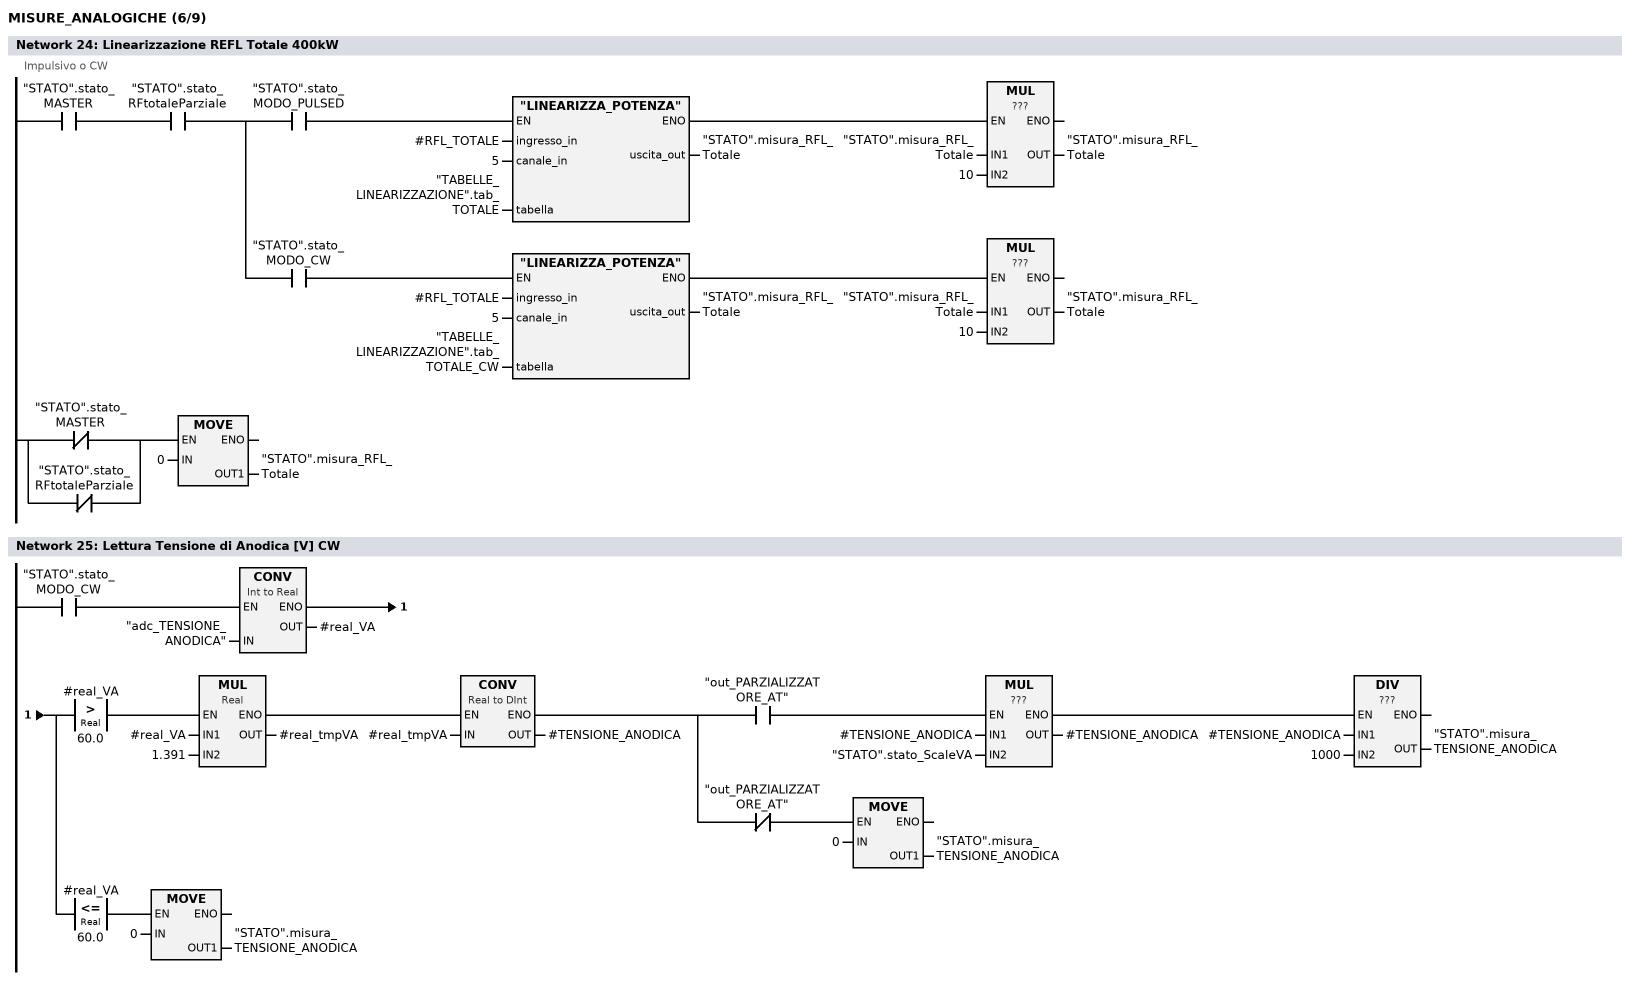
   RUNG wire#powerrail
      Contact( "STATO".stato_MASTER )
      Contact( "STATO".stato_RFtotaleParziale )
      wire#w1
      Contact( "STATO".stato_MODO_PULSED )
      "LINEARIZZA_POTENZA"(ingresso_in := #RFL_TOTALE, canale_in := 5, tabella := "TABELLE_LINEARIZZAZIONE".tab_TOTALE, uscita_out => "STATO".misura_RFL_Totale)
      { S7_Templates := "SrcType := ???" } Mul(in1 := "STATO".misura_RFL_Totale, in2 := 10, out => "STATO".misura_RFL_Totale)
   END_RUNG
   RUNG wire#w1
      Contact( "STATO".stato_MODO_CW )
      "LINEARIZZA_POTENZA"(ingresso_in := #RFL_TOTALE, canale_in := 5, tabella := "TABELLE_LINEARIZZAZIONE".tab_TOTALE_CW, uscita_out => "STATO".misura_RFL_Totale)
      { S7_Templates := "SrcType := ???" } Mul(in1 := "STATO".misura_RFL_Totale, in2 := 10, out => "STATO".misura_RFL_Totale)
   END_RUNG
   RUNG wire#powerrail
      I_Contact( "STATO".stato_MASTER )
      wire#w2
      Move(in := 0, out1 => "STATO".misura_RFL_Totale)
   END_RUNG
   RUNG wire#powerrail
      I_Contact( "STATO".stato_RFtotaleParziale )
   END_RUNG wire#w2
   // the same network as SCL:
   #_w1 := "STATO".stato_MASTER AND "STATO".stato_RFtotaleParziale;
   "LINEARIZZA_POTENZA"(EN := #_w1 AND "STATO".stato_MODO_PULSED,
                        ingresso_in := #RFL_TOTALE,
                        canale_in := 5,
                        tabella := "TABELLE_LINEARIZZAZIONE".tab_TOTALE,
                        uscita_out => "STATO".misura_RFL_Totale,
                        ENO => #_w2);
   IF #_w2 THEN "STATO".misura_RFL_Totale := "STATO".misura_RFL_Totale * 10; END_IF;
   "LINEARIZZA_POTENZA"(EN := #_w1 AND "STATO".stato_MODO_CW,
                        ingresso_in := #RFL_TOTALE,
                        canale_in := 5,
                        tabella := "TABELLE_LINEARIZZAZIONE".tab_TOTALE_CW,
                        uscita_out => "STATO".misura_RFL_Totale,
                        ENO => #_w3);
   IF #_w3 THEN "STATO".misura_RFL_Totale := "STATO".misura_RFL_Totale * 10; END_IF;
   IF NOT "STATO".stato_MASTER OR NOT "STATO".stato_RFtotaleParziale THEN
       "STATO".misura_RFL_Totale := 0;
   END_IF;
END_REGION

REGION Network 25: Lettura Tensione di Anodica [V] CW
   RUNG wire#powerrail
      Contact( "STATO".stato_MODO_CW )
      { S7_Templates := "[SrcType := Int, DestType := Real]" } Convert(in := "adc_TENSIONE_ANODICA", out => #real_VA)
      wire#w1
      { S7_Templates := "SrcType := Real" } GT_Contact(in1 := #real_VA, in2 := 60.0)
      { S7_Templates := "SrcType := Real" } Mul(in1 := #real_VA, in2 := 1.391, out => #real_tmpVA)
      { S7_Templates := "[SrcType := Real, DestType := DInt]" } Convert(in := #real_tmpVA, out => #TENSIONE_ANODICA)
      wire#w2
      Contact( "out_PARZIALIZZATORE_AT" )
      { S7_Templates := "SrcType := ???" } Mul(in1 := #TENSIONE_ANODICA, in2 := "STATO".stato_ScaleVA, out => #TENSIONE_ANODICA)
      { S7_Templates := "SrcType := ???" } Div(in1 := #TENSIONE_ANODICA, in2 := 1000, out => "STATO".misura_TENSIONE_ANODICA)
   END_RUNG
   RUNG wire#w2
      I_Contact( "out_PARZIALIZZATORE_AT" )
      Move(in := 0, out1 => "STATO".misura_TENSIONE_ANODICA)
   END_RUNG
   RUNG wire#w1
      { S7_Templates := "SrcType := Real" } LE_Contact(in1 := #real_VA, in2 := 60.0)
      Move(in := 0, out1 => "STATO".misura_TENSIONE_ANODICA)
   END_RUNG
   // the same network as SCL:
   IF "STATO".stato_MODO_CW THEN #real_VA := INT_TO_REAL("adc_TENSIONE_ANODICA"); END_IF;
   #_w1 := "STATO".stato_MODO_CW AND (#real_VA > 60.0);
   IF #_w1 THEN
       #real_tmpVA := #real_VA * 1.391;
       #TENSIONE_ANODICA := REAL_TO_DINT(#real_tmpVA);
   END_IF;
   IF #_w1 AND "out_PARZIALIZZATORE_AT" THEN
       #TENSIONE_ANODICA := #TENSIONE_ANODICA * "STATO".stato_ScaleVA;
       "STATO".misura_TENSIONE_ANODICA := #TENSIONE_ANODICA / 1000;
   END_IF;
   IF #_w1 AND NOT "out_PARZIALIZZATORE_AT" THEN "STATO".misura_TENSIONE_ANODICA := 0; END_IF;
   IF "STATO".stato_MODO_CW AND (#real_VA <= 60.0) THEN "STATO".misura_TENSIONE_ANODICA := 0; END_IF;
END_REGION

REGION Network 26: Lettura Tensione di Anodica [V] PULSED
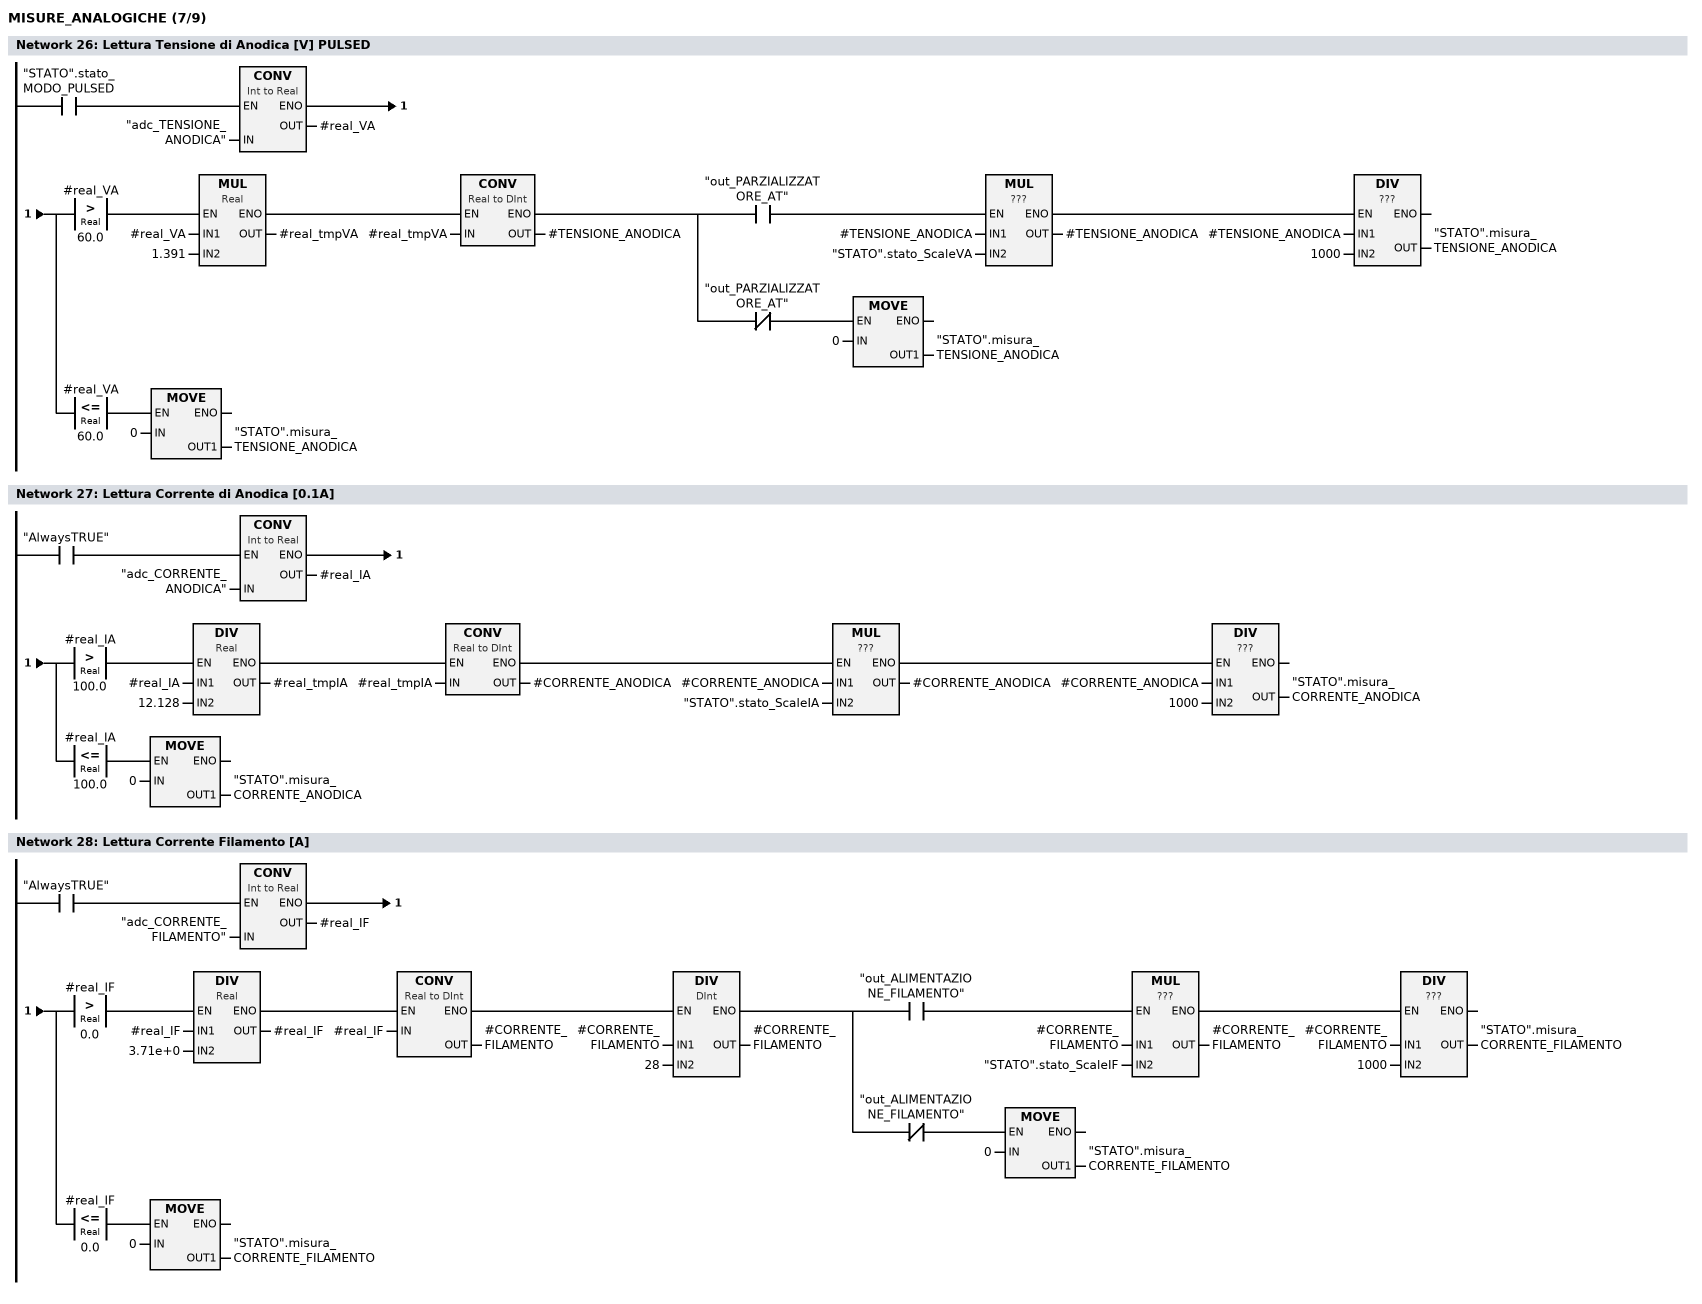
   RUNG wire#powerrail
      Contact( "STATO".stato_MODO_PULSED )
      { S7_Templates := "[SrcType := Int, DestType := Real]" } Convert(in := "adc_TENSIONE_ANODICA", out => #real_VA)
      wire#w1
      { S7_Templates := "SrcType := Real" } GT_Contact(in1 := #real_VA, in2 := 60.0)
      { S7_Templates := "SrcType := Real" } Mul(in1 := #real_VA, in2 := 1.391, out => #real_tmpVA)
      { S7_Templates := "[SrcType := Real, DestType := DInt]" } Convert(in := #real_tmpVA, out => #TENSIONE_ANODICA)
      wire#w2
      Contact( "out_PARZIALIZZATORE_AT" )
      { S7_Templates := "SrcType := ???" } Mul(in1 := #TENSIONE_ANODICA, in2 := "STATO".stato_ScaleVA, out => #TENSIONE_ANODICA)
      { S7_Templates := "SrcType := ???" } Div(in1 := #TENSIONE_ANODICA, in2 := 1000, out => "STATO".misura_TENSIONE_ANODICA)
   END_RUNG
   RUNG wire#w2
      I_Contact( "out_PARZIALIZZATORE_AT" )
      Move(in := 0, out1 => "STATO".misura_TENSIONE_ANODICA)
   END_RUNG
   RUNG wire#w1
      { S7_Templates := "SrcType := Real" } LE_Contact(in1 := #real_VA, in2 := 60.0)
      Move(in := 0, out1 => "STATO".misura_TENSIONE_ANODICA)
   END_RUNG
   // the same network as SCL:
   IF "STATO".stato_MODO_PULSED THEN #real_VA := INT_TO_REAL("adc_TENSIONE_ANODICA"); END_IF;
   #_w1 := "STATO".stato_MODO_PULSED AND (#real_VA > 60.0);
   IF #_w1 THEN
       #real_tmpVA := #real_VA * 1.391;
       #TENSIONE_ANODICA := REAL_TO_DINT(#real_tmpVA);
   END_IF;
   IF #_w1 AND "out_PARZIALIZZATORE_AT" THEN
       #TENSIONE_ANODICA := #TENSIONE_ANODICA * "STATO".stato_ScaleVA;
       "STATO".misura_TENSIONE_ANODICA := #TENSIONE_ANODICA / 1000;
   END_IF;
   IF #_w1 AND NOT "out_PARZIALIZZATORE_AT" THEN "STATO".misura_TENSIONE_ANODICA := 0; END_IF;
   IF "STATO".stato_MODO_PULSED AND (#real_VA <= 60.0) THEN "STATO".misura_TENSIONE_ANODICA := 0; END_IF;
END_REGION

REGION Network 27: Lettura Corrente di Anodica [0.1A]
   RUNG wire#powerrail
      Contact( "AlwaysTRUE" )
      { S7_Templates := "[SrcType := Int, DestType := Real]" } Convert(in := "adc_CORRENTE_ANODICA", out => #real_IA)
      wire#w1
      { S7_Templates := "SrcType := Real" } GT_Contact(in1 := #real_IA, in2 := 100.0)
      { S7_Templates := "SrcType := Real" } Div(in1 := #real_IA, in2 := 12.128, out => #real_tmpIA)
      { S7_Templates := "[SrcType := Real, DestType := DInt]" } Convert(in := #real_tmpIA, out => #CORRENTE_ANODICA)
      { S7_Templates := "SrcType := ???" } Mul(in1 := #CORRENTE_ANODICA, in2 := "STATO".stato_ScaleIA, out => #CORRENTE_ANODICA)
      { S7_Templates := "SrcType := ???" } Div(in1 := #CORRENTE_ANODICA, in2 := 1000, out => "STATO".misura_CORRENTE_ANODICA)
   END_RUNG
   RUNG wire#w1
      { S7_Templates := "SrcType := Real" } LE_Contact(in1 := #real_IA, in2 := 100.0)
      Move(in := 0, out1 => "STATO".misura_CORRENTE_ANODICA)
   END_RUNG
   // the same network as SCL:
   IF "AlwaysTRUE" THEN #real_IA := INT_TO_REAL("adc_CORRENTE_ANODICA"); END_IF;
   IF "AlwaysTRUE" AND (#real_IA > 100.0) THEN
       #real_tmpIA := #real_IA / 12.128;
       #CORRENTE_ANODICA := REAL_TO_DINT(#real_tmpIA);
       #CORRENTE_ANODICA := #CORRENTE_ANODICA * "STATO".stato_ScaleIA;
       "STATO".misura_CORRENTE_ANODICA := #CORRENTE_ANODICA / 1000;
   END_IF;
   IF "AlwaysTRUE" AND (#real_IA <= 100.0) THEN "STATO".misura_CORRENTE_ANODICA := 0; END_IF;
END_REGION

REGION Network 28: Lettura Corrente Filamento [A]
   RUNG wire#powerrail
      Contact( "AlwaysTRUE" )
      { S7_Templates := "[SrcType := Int, DestType := Real]" } Convert(in := "adc_CORRENTE_FILAMENTO", out => #real_IF)
      wire#w1
      { S7_Templates := "SrcType := Real" } GT_Contact(in1 := #real_IF, in2 := 0.0)
      { S7_Templates := "SrcType := Real" } Div(in1 := #real_IF, in2 := 3.71e+0, out => #real_IF)
      { S7_Templates := "[SrcType := Real, DestType := DInt]" } Convert(in := #real_IF, out => #CORRENTE_FILAMENTO)
      { S7_Templates := "SrcType := DInt" } Div(in1 := #CORRENTE_FILAMENTO, in2 := 28, out => #CORRENTE_FILAMENTO)
      wire#w2
      Contact( "out_ALIMENTAZIONE_FILAMENTO" )
      { S7_Templates := "SrcType := ???" } Mul(in1 := #CORRENTE_FILAMENTO, in2 := "STATO".stato_ScaleIF, out => #CORRENTE_FILAMENTO)
      { S7_Templates := "SrcType := ???" } Div(in1 := #CORRENTE_FILAMENTO, in2 := 1000, out => "STATO".misura_CORRENTE_FILAMENTO)
   END_RUNG
   RUNG wire#w2
      I_Contact( "out_ALIMENTAZIONE_FILAMENTO" )
      Move(in := 0, out1 => "STATO".misura_CORRENTE_FILAMENTO)
   END_RUNG
   RUNG wire#w1
      { S7_Templates := "SrcType := Real" } LE_Contact(in1 := #real_IF, in2 := 0.0)
      Move(in := 0, out1 => "STATO".misura_CORRENTE_FILAMENTO)
   END_RUNG
   // the same network as SCL:
   IF "AlwaysTRUE" THEN #real_IF := INT_TO_REAL("adc_CORRENTE_FILAMENTO"); END_IF;
   #_w1 := "AlwaysTRUE" AND (#real_IF > 0.0);
   IF #_w1 THEN
       #real_IF := #real_IF / 3.71e+0;
       #CORRENTE_FILAMENTO := REAL_TO_DINT(#real_IF);
       #CORRENTE_FILAMENTO := #CORRENTE_FILAMENTO / 28;
   END_IF;
   IF #_w1 AND "out_ALIMENTAZIONE_FILAMENTO" THEN
       #CORRENTE_FILAMENTO := #CORRENTE_FILAMENTO * "STATO".stato_ScaleIF;
       "STATO".misura_CORRENTE_FILAMENTO := #CORRENTE_FILAMENTO / 1000;
   END_IF;
   IF #_w1 AND NOT "out_ALIMENTAZIONE_FILAMENTO" THEN "STATO".misura_CORRENTE_FILAMENTO := 0; END_IF;
   IF "AlwaysTRUE" AND (#real_IF <= 0.0) THEN "STATO".misura_CORRENTE_FILAMENTO := 0; END_IF;
END_REGION

REGION Network 29: Lettura Tensione VG1 [V]
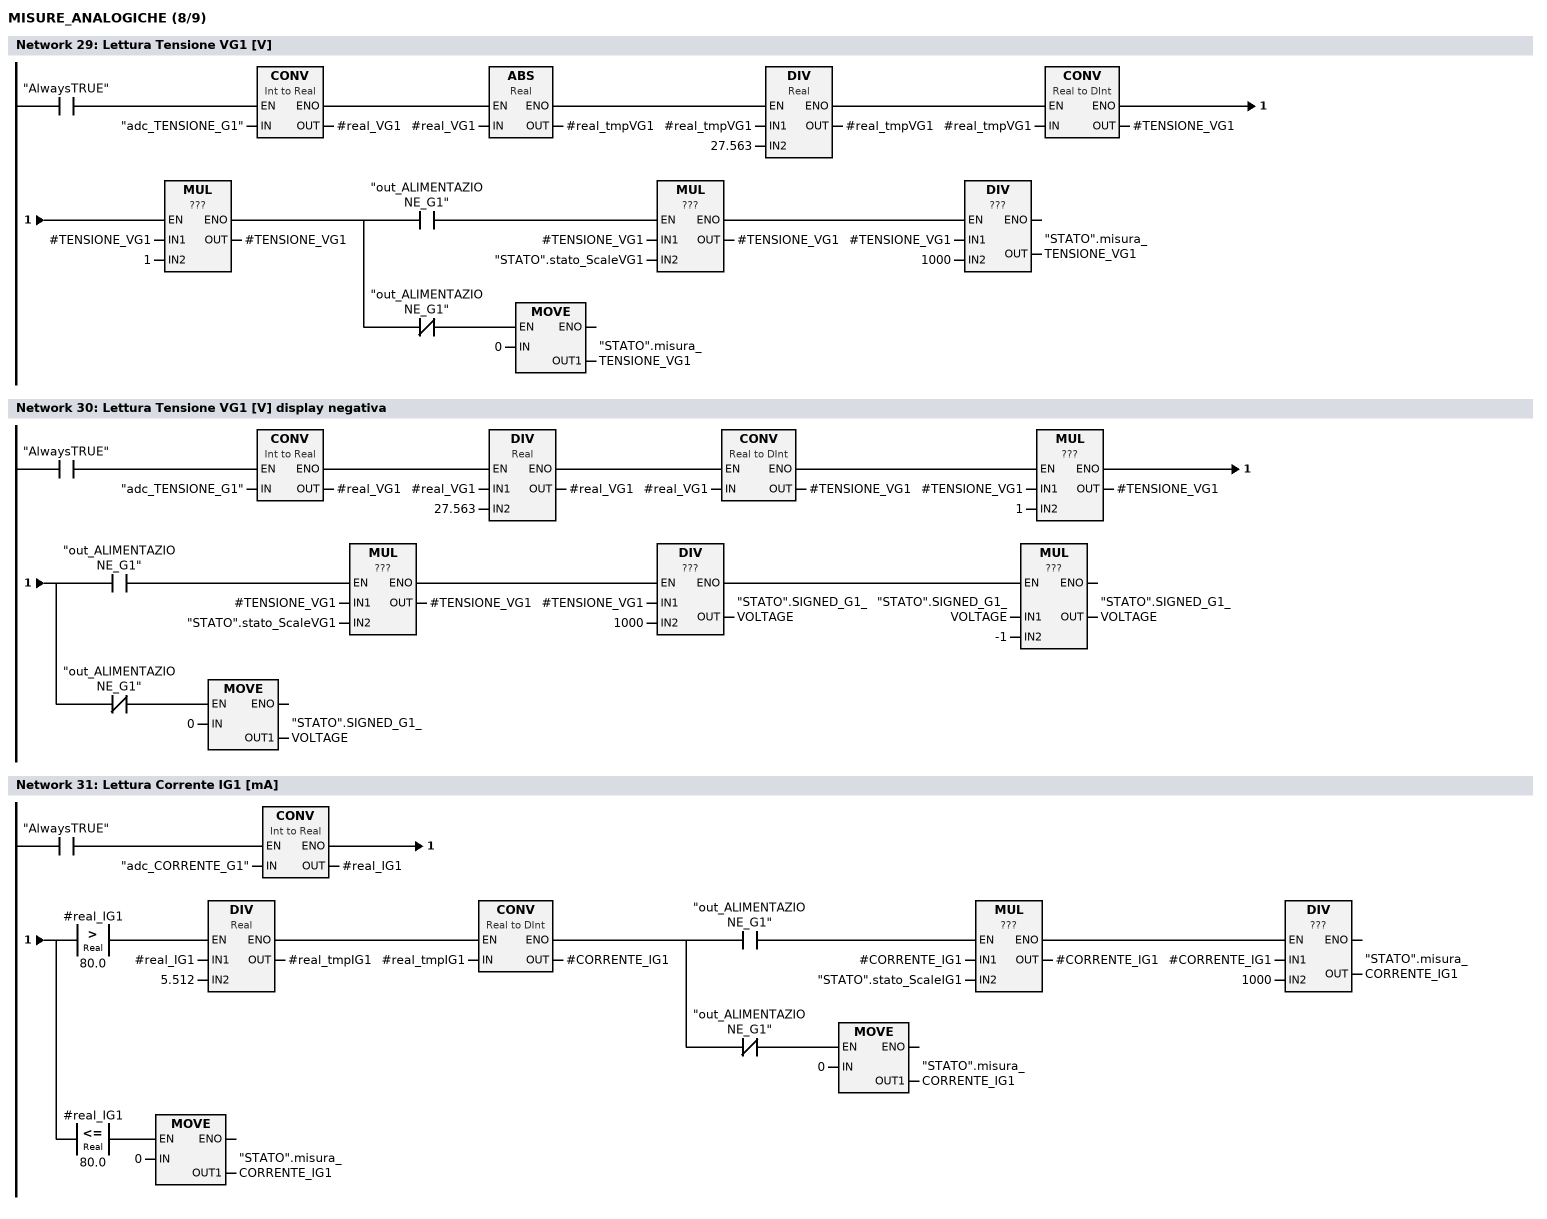
   RUNG wire#powerrail
      Contact( "AlwaysTRUE" )
      { S7_Templates := "[SrcType := Int, DestType := Real]" } Convert(in := "adc_TENSIONE_G1", out => #real_VG1)
      { S7_Templates := "SrcType := Real" } Abs(in := #real_VG1, out => #real_tmpVG1)
      { S7_Templates := "SrcType := Real" } Div(in1 := #real_tmpVG1, in2 := 27.563, out => #real_tmpVG1)
      { S7_Templates := "[SrcType := Real, DestType := DInt]" } Convert(in := #real_tmpVG1, out => #TENSIONE_VG1)
      { S7_Templates := "SrcType := ???" } Mul(in1 := #TENSIONE_VG1, in2 := 1, out => #TENSIONE_VG1)
      wire#w1
      Contact( "out_ALIMENTAZIONE_G1" )
      { S7_Templates := "SrcType := ???" } Mul(in1 := #TENSIONE_VG1, in2 := "STATO".stato_ScaleVG1, out => #TENSIONE_VG1)
      { S7_Templates := "SrcType := ???" } Div(in1 := #TENSIONE_VG1, in2 := 1000, out => "STATO".misura_TENSIONE_VG1)
   END_RUNG
   RUNG wire#w1
      I_Contact( "out_ALIMENTAZIONE_G1" )
      Move(in := 0, out1 => "STATO".misura_TENSIONE_VG1)
   END_RUNG
   // the same network as SCL:
   IF "AlwaysTRUE" THEN
       #real_VG1 := INT_TO_REAL("adc_TENSIONE_G1");
       #real_tmpVG1 := ABS(#real_VG1);
       #real_tmpVG1 := #real_tmpVG1 / 27.563;
       #TENSIONE_VG1 := REAL_TO_DINT(#real_tmpVG1);
       #TENSIONE_VG1 := #TENSIONE_VG1 * 1;
   END_IF;
   IF "AlwaysTRUE" AND "out_ALIMENTAZIONE_G1" THEN
       #TENSIONE_VG1 := #TENSIONE_VG1 * "STATO".stato_ScaleVG1;
       "STATO".misura_TENSIONE_VG1 := #TENSIONE_VG1 / 1000;
   END_IF;
   IF "AlwaysTRUE" AND NOT "out_ALIMENTAZIONE_G1" THEN "STATO".misura_TENSIONE_VG1 := 0; END_IF;
END_REGION

REGION Network 30: Lettura Tensione VG1 [V] display negativa
   RUNG wire#powerrail
      Contact( "AlwaysTRUE" )
      { S7_Templates := "[SrcType := Int, DestType := Real]" } Convert(in := "adc_TENSIONE_G1", out => #real_VG1)
      { S7_Templates := "SrcType := Real" } Div(in1 := #real_VG1, in2 := 27.563, out => #real_VG1)
      { S7_Templates := "[SrcType := Real, DestType := DInt]" } Convert(in := #real_VG1, out => #TENSIONE_VG1)
      { S7_Templates := "SrcType := ???" } Mul(in1 := #TENSIONE_VG1, in2 := 1, out => #TENSIONE_VG1)
      wire#w1
      Contact( "out_ALIMENTAZIONE_G1" )
      { S7_Templates := "SrcType := ???" } Mul(in1 := #TENSIONE_VG1, in2 := "STATO".stato_ScaleVG1, out => #TENSIONE_VG1)
      { S7_Templates := "SrcType := ???" } Div(in1 := #TENSIONE_VG1, in2 := 1000, out => "STATO".SIGNED_G1_VOLTAGE)
      { S7_Templates := "SrcType := ???" } Mul(in1 := "STATO".SIGNED_G1_VOLTAGE, in2 := -1, out => "STATO".SIGNED_G1_VOLTAGE)
   END_RUNG
   RUNG wire#w1
      I_Contact( "out_ALIMENTAZIONE_G1" )
      Move(in := 0, out1 => "STATO".SIGNED_G1_VOLTAGE)
   END_RUNG
   // the same network as SCL:
   IF "AlwaysTRUE" THEN
       #real_VG1 := INT_TO_REAL("adc_TENSIONE_G1");
       #real_VG1 := #real_VG1 / 27.563;
       #TENSIONE_VG1 := REAL_TO_DINT(#real_VG1);
       #TENSIONE_VG1 := #TENSIONE_VG1 * 1;
   END_IF;
   IF "AlwaysTRUE" AND "out_ALIMENTAZIONE_G1" THEN
       #TENSIONE_VG1 := #TENSIONE_VG1 * "STATO".stato_ScaleVG1;
       "STATO".SIGNED_G1_VOLTAGE := #TENSIONE_VG1 / 1000;
       "STATO".SIGNED_G1_VOLTAGE := "STATO".SIGNED_G1_VOLTAGE * (-1);
   END_IF;
   IF "AlwaysTRUE" AND NOT "out_ALIMENTAZIONE_G1" THEN "STATO".SIGNED_G1_VOLTAGE := 0; END_IF;
END_REGION

REGION Network 31: Lettura Corrente IG1 [mA]
   RUNG wire#powerrail
      Contact( "AlwaysTRUE" )
      { S7_Templates := "[SrcType := Int, DestType := Real]" } Convert(in := "adc_CORRENTE_G1", out => #real_IG1)
      wire#w1
      { S7_Templates := "SrcType := Real" } GT_Contact(in1 := #real_IG1, in2 := 80.0)
      { S7_Templates := "SrcType := Real" } Div(in1 := #real_IG1, in2 := 5.512, out => #real_tmpIG1)
      { S7_Templates := "[SrcType := Real, DestType := DInt]" } Convert(in := #real_tmpIG1, out => #CORRENTE_IG1)
      wire#w2
      Contact( "out_ALIMENTAZIONE_G1" )
      { S7_Templates := "SrcType := ???" } Mul(in1 := #CORRENTE_IG1, in2 := "STATO".stato_ScaleIG1, out => #CORRENTE_IG1)
      { S7_Templates := "SrcType := ???" } Div(in1 := #CORRENTE_IG1, in2 := 1000, out => "STATO".misura_CORRENTE_IG1)
   END_RUNG
   RUNG wire#w2
      I_Contact( "out_ALIMENTAZIONE_G1" )
      Move(in := 0, out1 => "STATO".misura_CORRENTE_IG1)
   END_RUNG
   RUNG wire#w1
      { S7_Templates := "SrcType := Real" } LE_Contact(in1 := #real_IG1, in2 := 80.0)
      Move(in := 0, out1 => "STATO".misura_CORRENTE_IG1)
   END_RUNG
   // the same network as SCL:
   IF "AlwaysTRUE" THEN #real_IG1 := INT_TO_REAL("adc_CORRENTE_G1"); END_IF;
   #_w1 := "AlwaysTRUE" AND (#real_IG1 > 80.0);
   IF #_w1 THEN
       #real_tmpIG1 := #real_IG1 / 5.512;
       #CORRENTE_IG1 := REAL_TO_DINT(#real_tmpIG1);
   END_IF;
   IF #_w1 AND "out_ALIMENTAZIONE_G1" THEN
       #CORRENTE_IG1 := #CORRENTE_IG1 * "STATO".stato_ScaleIG1;
       "STATO".misura_CORRENTE_IG1 := #CORRENTE_IG1 / 1000;
   END_IF;
   IF #_w1 AND NOT "out_ALIMENTAZIONE_G1" THEN "STATO".misura_CORRENTE_IG1 := 0; END_IF;
   IF "AlwaysTRUE" AND (#real_IG1 <= 80.0) THEN "STATO".misura_CORRENTE_IG1 := 0; END_IF;
END_REGION

REGION Network 32: Lettura Tensione VG2 [V]
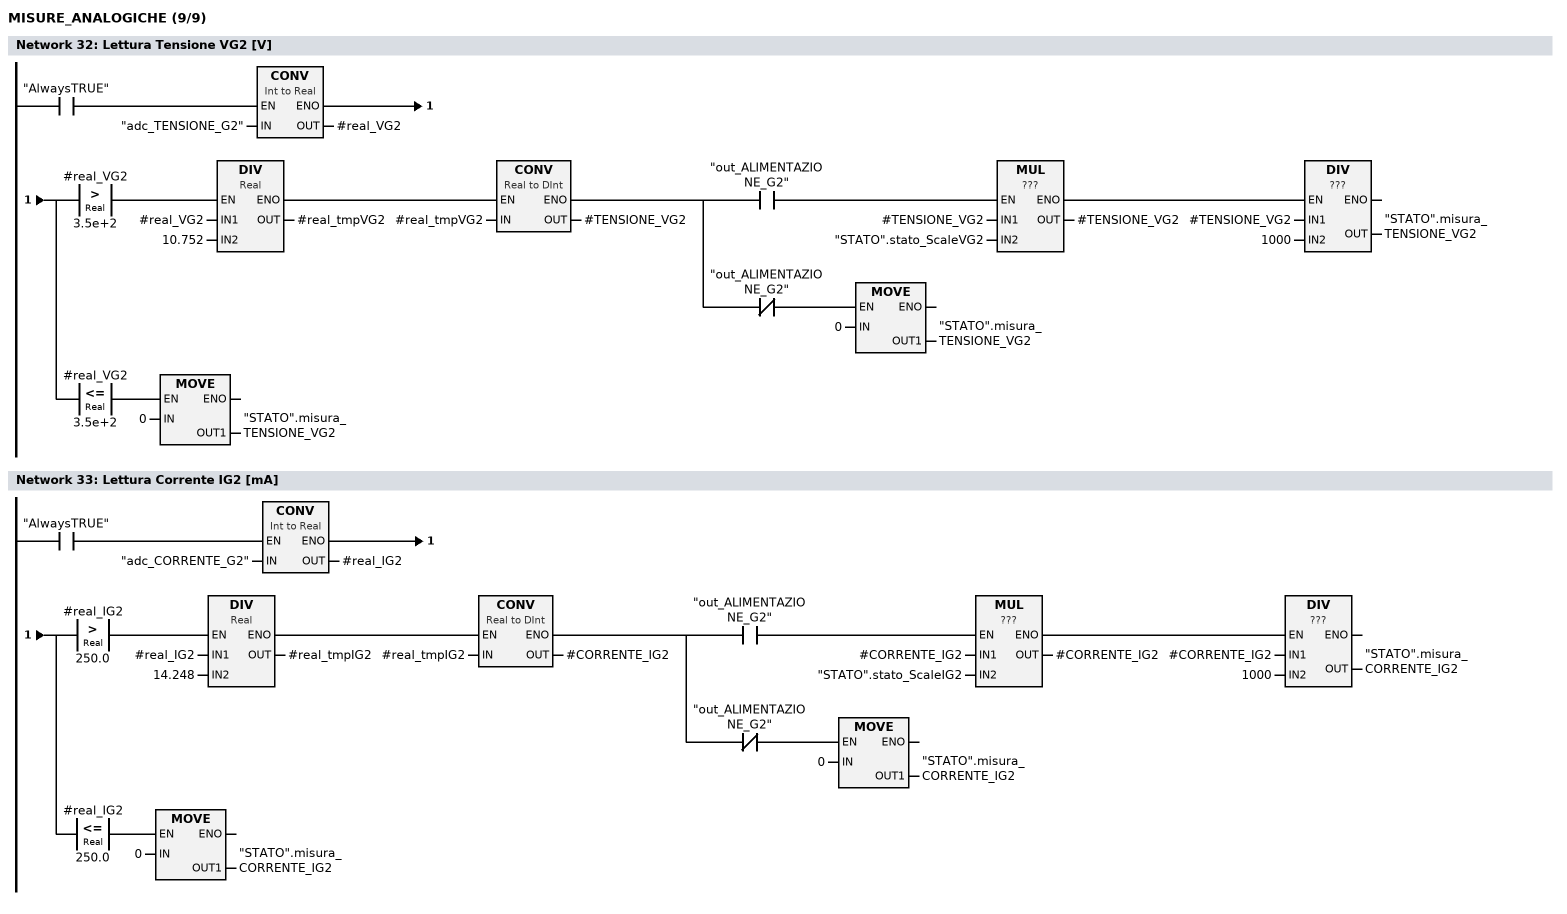
   RUNG wire#powerrail
      Contact( "AlwaysTRUE" )
      { S7_Templates := "[SrcType := Int, DestType := Real]" } Convert(in := "adc_TENSIONE_G2", out => #real_VG2)
      wire#w1
      { S7_Templates := "SrcType := Real" } GT_Contact(in1 := #real_VG2, in2 := 3.5e+2)
      { S7_Templates := "SrcType := Real" } Div(in1 := #real_VG2, in2 := 10.752, out => #real_tmpVG2)
      { S7_Templates := "[SrcType := Real, DestType := DInt]" } Convert(in := #real_tmpVG2, out => #TENSIONE_VG2)
      wire#w2
      Contact( "out_ALIMENTAZIONE_G2" )
      { S7_Templates := "SrcType := ???" } Mul(in1 := #TENSIONE_VG2, in2 := "STATO".stato_ScaleVG2, out => #TENSIONE_VG2)
      { S7_Templates := "SrcType := ???" } Div(in1 := #TENSIONE_VG2, in2 := 1000, out => "STATO".misura_TENSIONE_VG2)
   END_RUNG
   RUNG wire#w2
      I_Contact( "out_ALIMENTAZIONE_G2" )
      Move(in := 0, out1 => "STATO".misura_TENSIONE_VG2)
   END_RUNG
   RUNG wire#w1
      { S7_Templates := "SrcType := Real" } LE_Contact(in1 := #real_VG2, in2 := 3.5e+2)
      Move(in := 0, out1 => "STATO".misura_TENSIONE_VG2)
   END_RUNG
   // the same network as SCL:
   IF "AlwaysTRUE" THEN #real_VG2 := INT_TO_REAL("adc_TENSIONE_G2"); END_IF;
   #_w1 := "AlwaysTRUE" AND (#real_VG2 > 3.5e+2);
   IF #_w1 THEN
       #real_tmpVG2 := #real_VG2 / 10.752;
       #TENSIONE_VG2 := REAL_TO_DINT(#real_tmpVG2);
   END_IF;
   IF #_w1 AND "out_ALIMENTAZIONE_G2" THEN
       #TENSIONE_VG2 := #TENSIONE_VG2 * "STATO".stato_ScaleVG2;
       "STATO".misura_TENSIONE_VG2 := #TENSIONE_VG2 / 1000;
   END_IF;
   IF #_w1 AND NOT "out_ALIMENTAZIONE_G2" THEN "STATO".misura_TENSIONE_VG2 := 0; END_IF;
   IF "AlwaysTRUE" AND (#real_VG2 <= 3.5e+2) THEN "STATO".misura_TENSIONE_VG2 := 0; END_IF;
END_REGION

REGION Network 33: Lettura Corrente IG2 [mA]
   RUNG wire#powerrail
      Contact( "AlwaysTRUE" )
      { S7_Templates := "[SrcType := Int, DestType := Real]" } Convert(in := "adc_CORRENTE_G2", out => #real_IG2)
      wire#w1
      { S7_Templates := "SrcType := Real" } GT_Contact(in1 := #real_IG2, in2 := 250.0)
      { S7_Templates := "SrcType := Real" } Div(in1 := #real_IG2, in2 := 14.248, out => #real_tmpIG2)
      { S7_Templates := "[SrcType := Real, DestType := DInt]" } Convert(in := #real_tmpIG2, out => #CORRENTE_IG2)
      wire#w2
      Contact( "out_ALIMENTAZIONE_G2" )
      { S7_Templates := "SrcType := ???" } Mul(in1 := #CORRENTE_IG2, in2 := "STATO".stato_ScaleIG2, out => #CORRENTE_IG2)
      { S7_Templates := "SrcType := ???" } Div(in1 := #CORRENTE_IG2, in2 := 1000, out => "STATO".misura_CORRENTE_IG2)
   END_RUNG
   RUNG wire#w2
      I_Contact( "out_ALIMENTAZIONE_G2" )
      Move(in := 0, out1 => "STATO".misura_CORRENTE_IG2)
   END_RUNG
   RUNG wire#w1
      { S7_Templates := "SrcType := Real" } LE_Contact(in1 := #real_IG2, in2 := 250.0)
      Move(in := 0, out1 => "STATO".misura_CORRENTE_IG2)
   END_RUNG
   // the same network as SCL:
   IF "AlwaysTRUE" THEN #real_IG2 := INT_TO_REAL("adc_CORRENTE_G2"); END_IF;
   #_w1 := "AlwaysTRUE" AND (#real_IG2 > 250.0);
   IF #_w1 THEN
       #real_tmpIG2 := #real_IG2 / 14.248;
       #CORRENTE_IG2 := REAL_TO_DINT(#real_tmpIG2);
   END_IF;
   IF #_w1 AND "out_ALIMENTAZIONE_G2" THEN
       #CORRENTE_IG2 := #CORRENTE_IG2 * "STATO".stato_ScaleIG2;
       "STATO".misura_CORRENTE_IG2 := #CORRENTE_IG2 / 1000;
   END_IF;
   IF #_w1 AND NOT "out_ALIMENTAZIONE_G2" THEN "STATO".misura_CORRENTE_IG2 := 0; END_IF;
   IF "AlwaysTRUE" AND (#real_IG2 <= 250.0) THEN "STATO".misura_CORRENTE_IG2 := 0; END_IF;
END_REGION
END_FUNCTION

FUNCTION "REGOLA_ANODICA" : Void   // FC2, LAD
{ S7_Optimized_Access := 'FALSE' }
VERSION : 0.1
   VAR_TEMP   // added for the SCL form of the ladder/FBD networks
      _w1 : Bool;
   END_VAR
BEGIN

REGION Network 1
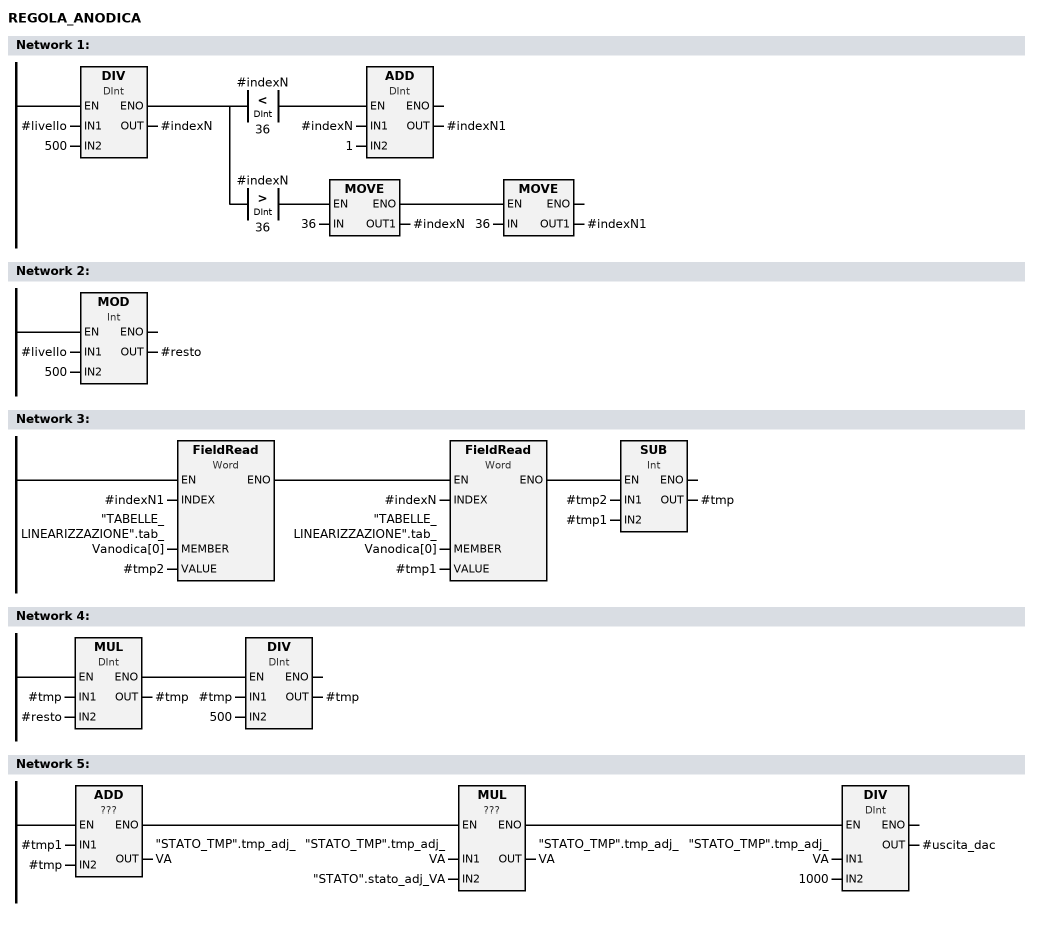
   RUNG wire#powerrail
      { S7_Templates := "SrcType := DInt" } Div(in1 := #livello, in2 := 500, out => #indexN)
      wire#w1
      { S7_Templates := "SrcType := DInt" } LT_Contact(in1 := #indexN, in2 := 36)
      { S7_Templates := "SrcType := DInt" } Add(in1 := #indexN, in2 := 1, out => #indexN1)
   END_RUNG
   RUNG wire#w1
      { S7_Templates := "SrcType := DInt" } GT_Contact(in1 := #indexN, in2 := 36)
      Move(in := 36, out1 => #indexN)
      Move(in := 36, out1 => #indexN1)
   END_RUNG
   // the same network as SCL:
   #indexN := #livello / 500;
   IF #indexN < 36 THEN #indexN1 := #indexN + 1; END_IF;
   #_w1 := #indexN > 36;
   IF #_w1 THEN
       #indexN := 36;
       #indexN1 := 36;
   END_IF;
END_REGION

REGION Network 2
   RUNG wire#powerrail
      { S7_Templates := "SrcType := Int" } Mod(in1 := #livello, in2 := 500, out => #resto)
   END_RUNG
   // the same network as SCL:
   #resto := #livello MOD 500;
END_REGION

REGION Network 3
   // no SCL statement known for FieldRead: written as a call
   // ENO of a box is taken as its EN; it also drops when the box reports an error
   FieldRead(index := #indexN1, member := "TABELLE_LINEARIZZAZIONE".tab_Vanodica[0], value := #tmp2);
   FieldRead(index := #indexN, member := "TABELLE_LINEARIZZAZIONE".tab_Vanodica[0], value := #tmp1);
   #tmp := #tmp2 - #tmp1;
END_REGION

REGION Network 4
   RUNG wire#powerrail
      { S7_Templates := "SrcType := DInt" } Mul(in1 := #tmp, in2 := #resto, out => #tmp)
      { S7_Templates := "SrcType := DInt" } Div(in1 := #tmp, in2 := 500, out => #tmp)
   END_RUNG
   // the same network as SCL:
   #tmp := #tmp * #resto;
   #tmp := #tmp / 500;
END_REGION

REGION Network 5
   RUNG wire#powerrail
      { S7_Templates := "SrcType := ???" } Add(in1 := #tmp1, in2 := #tmp, out => "STATO_TMP".tmp_adj_VA)
      { S7_Templates := "SrcType := ???" } Mul(in1 := "STATO_TMP".tmp_adj_VA, in2 := "STATO".stato_adj_VA, out => "STATO_TMP".tmp_adj_VA)
      { S7_Templates := "SrcType := DInt" } Div(in1 := "STATO_TMP".tmp_adj_VA, in2 := 1000, out => #uscita_dac)
   END_RUNG
   // the same network as SCL:
   "STATO_TMP".tmp_adj_VA := #tmp1 + #tmp;
   "STATO_TMP".tmp_adj_VA := "STATO_TMP".tmp_adj_VA * "STATO".stato_adj_VA;
   #uscita_dac := "STATO_TMP".tmp_adj_VA / 1000;
END_REGION
END_FUNCTION

FUNCTION "SERIAL_SEND" : Void   // FC3, LAD
TITLE = SERIAL_SEND
{ S7_Optimized_Access := 'FALSE' }
VERSION : 0.1
// In questa Function Block preparo il messaggio da inviare discriminandone il tipo.
   VAR_TEMP   // added for the SCL form of the ladder/FBD networks
      _w1 : Bool;
   END_VAR
BEGIN

REGION Network 1: Ho finito il giro delle richieste di stato
   // Riparto con le richieste di stato dal primo slave.
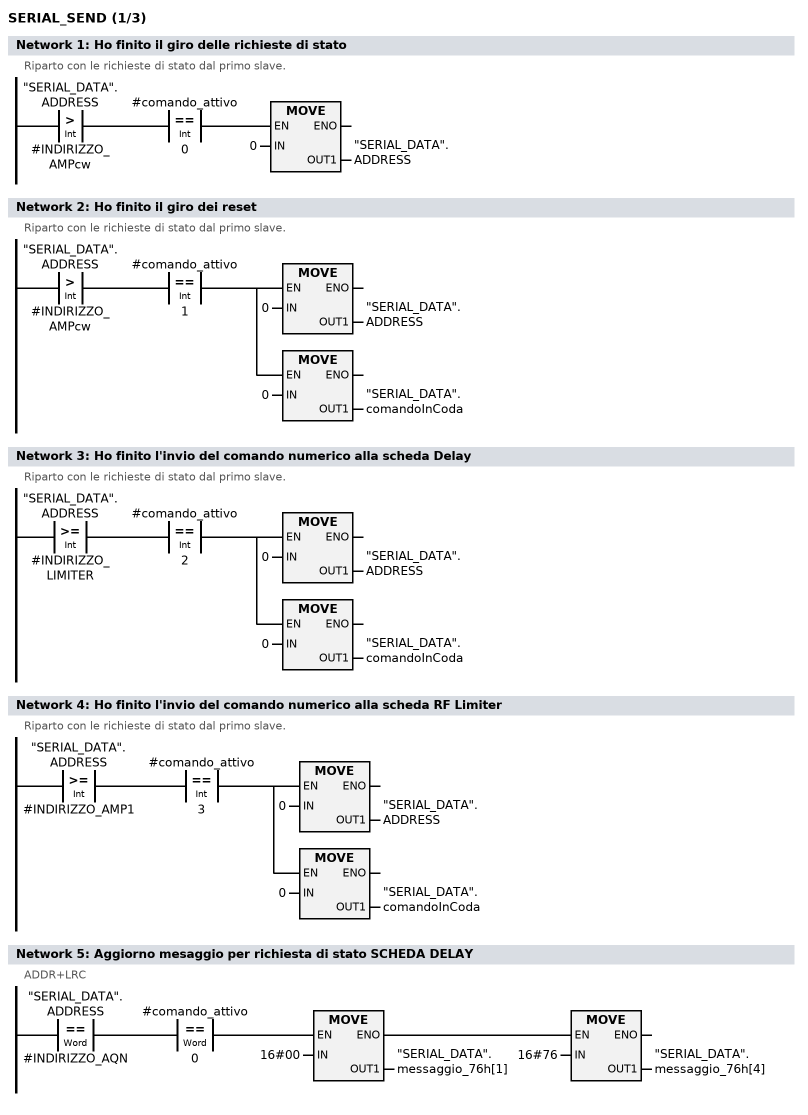
   RUNG wire#powerrail
      { S7_Templates := "SrcType := Int" } GT_Contact(in1 := "SERIAL_DATA".ADDRESS, in2 := #INDIRIZZO_AMPcw)
      { S7_Templates := "SrcType := Int" } EQ_Contact(in1 := #comando_attivo, in2 := 0)
      Move(in := 0, out1 => "SERIAL_DATA".ADDRESS)
   END_RUNG
   // the same network as SCL:
   IF ("SERIAL_DATA".ADDRESS > #INDIRIZZO_AMPcw) AND (#comando_attivo = 0) THEN
       "SERIAL_DATA".ADDRESS := 0;
   END_IF;
END_REGION

REGION Network 2: Ho finito il giro dei reset
   // Riparto con le richieste di stato dal primo slave.
   RUNG wire#powerrail
      { S7_Templates := "SrcType := Int" } GT_Contact(in1 := "SERIAL_DATA".ADDRESS, in2 := #INDIRIZZO_AMPcw)
      { S7_Templates := "SrcType := Int" } EQ_Contact(in1 := #comando_attivo, in2 := 1)
      wire#w1
      Move(in := 0, out1 => "SERIAL_DATA".ADDRESS)
   END_RUNG
   RUNG wire#w1
      Move(in := 0, out1 => "SERIAL_DATA".comandoInCoda)
   END_RUNG
   // the same network as SCL:
   #_w1 := ("SERIAL_DATA".ADDRESS > #INDIRIZZO_AMPcw) AND (#comando_attivo = 1);
   IF #_w1 THEN
       "SERIAL_DATA".ADDRESS := 0;
       "SERIAL_DATA".comandoInCoda := 0;
   END_IF;
END_REGION

REGION Network 3: Ho finito l'invio del comando numerico alla scheda Delay
   // Riparto con le richieste di stato dal primo slave.
   RUNG wire#powerrail
      { S7_Templates := "SrcType := Int" } GE_Contact(in1 := "SERIAL_DATA".ADDRESS, in2 := #INDIRIZZO_LIMITER)
      { S7_Templates := "SrcType := Int" } EQ_Contact(in1 := #comando_attivo, in2 := 2)
      wire#w1
      Move(in := 0, out1 => "SERIAL_DATA".ADDRESS)
   END_RUNG
   RUNG wire#w1
      Move(in := 0, out1 => "SERIAL_DATA".comandoInCoda)
   END_RUNG
   // the same network as SCL:
   #_w1 := ("SERIAL_DATA".ADDRESS >= #INDIRIZZO_LIMITER) AND (#comando_attivo = 2);
   IF #_w1 THEN
       "SERIAL_DATA".ADDRESS := 0;
       "SERIAL_DATA".comandoInCoda := 0;
   END_IF;
END_REGION

REGION Network 4: Ho finito l'invio del comando numerico alla scheda RF Limiter
   // Riparto con le richieste di stato dal primo slave.
   RUNG wire#powerrail
      { S7_Templates := "SrcType := Int" } GE_Contact(in1 := "SERIAL_DATA".ADDRESS, in2 := #INDIRIZZO_AMP1)
      { S7_Templates := "SrcType := Int" } EQ_Contact(in1 := #comando_attivo, in2 := 3)
      wire#w1
      Move(in := 0, out1 => "SERIAL_DATA".ADDRESS)
   END_RUNG
   RUNG wire#w1
      Move(in := 0, out1 => "SERIAL_DATA".comandoInCoda)
   END_RUNG
   // the same network as SCL:
   #_w1 := ("SERIAL_DATA".ADDRESS >= #INDIRIZZO_AMP1) AND (#comando_attivo = 3);
   IF #_w1 THEN
       "SERIAL_DATA".ADDRESS := 0;
       "SERIAL_DATA".comandoInCoda := 0;
   END_IF;
END_REGION

REGION Network 5: Aggiorno mesaggio per richiesta di stato SCHEDA DELAY
   // ADDR+LRC
   RUNG wire#powerrail
      { S7_Templates := "SrcType := Word" } EQ_Contact(in1 := "SERIAL_DATA".ADDRESS, in2 := #INDIRIZZO_AQN)
      { S7_Templates := "SrcType := Word" } EQ_Contact(in1 := #comando_attivo, in2 := 0)
      Move(in := 16#00, out1 => "SERIAL_DATA".messaggio_76h[1])
      Move(in := 16#76, out1 => "SERIAL_DATA".messaggio_76h[4])
   END_RUNG
   // the same network as SCL:
   IF ("SERIAL_DATA".ADDRESS = #INDIRIZZO_AQN) AND (#comando_attivo = 0) THEN
       "SERIAL_DATA".messaggio_76h[1] := 16#00;
       "SERIAL_DATA".messaggio_76h[4] := 16#76;
   END_IF;
END_REGION

